   "Tank 5S Tank Vent Valve 2 Feedback - Closed" : Bool = PLC "Tank 5S Tank Vent Valve 2 Feedback - Closed" AT %I54.5, 1 s
   "RIO5_SPR_DI_54_6" : Bool = PLC RIO5_SPR_DI_54_6 AT %I54.6, 1 s
   "RIO5_SPR_DI_54_7" : Bool = PLC RIO5_SPR_DI_54_7 AT %I54.7, 1 s
   "Tank 5P BWT Level High High Switch" : Bool = PLC "Tank 5P BWT Level High High Switch" AT %I57.0, 1 s
   "RIO5 Tanks Pressure Switch Hi Hi" : Bool = PLC "RIO5 Tanks Pressure Switch Hi Hi" AT %I57.1, 1 s
   "Tank 5S BWT Level High High Switch" : Bool = PLC "Tank 5S BWT Level High High Switch" AT %I57.2, 1 s
   "RIO5_SPR_DI_57_3" : Bool = PLC RIO5_SPR_DI_57_3 AT %I57.3, 1 s
   "RIO5_SPR_DI_57_4" : Bool = PLC RIO5_SPR_DI_57_4 AT %I57.4, 1 s
   "RIO5_SPR_DI_57_5" : Bool = PLC RIO5_SPR_DI_57_5 AT %I57.5, 1 s
   "RIO5_SPR_DI_57_6" : Bool = PLC RIO5_SPR_DI_57_6 AT %I57.6, 1 s
   "RIO5_SPR_DI_57_7" : Bool = PLC RIO5_SPR_DI_57_7 AT %I57.7, 1 s
   "Tank 6P GTT Isolation Valve Feedback - Opened" : Bool = PLC "Tank 6P GTT Isolation Valve Feedback - Opened" AT %I60.0, 1 s
   "Tank 6P GTT Isolation Valve Feedback - Closed" : Bool = PLC "Tank 6P GTT Isolation Valve Feedback - Closed" AT %I60.1, 1 s
   "Tank 6P Tank Vent Valve 1 Feedback - Opened" : Bool = PLC "Tank 6P Tank Vent Valve 1 Feedback - Opened" AT %I60.2, 1 s
   "Tank 6P Tank Vent Valve 1 Feedback - Closed" : Bool = PLC "Tank 6P Tank Vent Valve 1 Feedback - Closed" AT %I60.3, 1 s
   "Tank 6P Tank Vent Valve 2 Feedback - Opened" : Bool = PLC "Tank 6P Tank Vent Valve 2 Feedback - Opened" AT %I60.4, 1 s
   "Tank 6P Tank Vent Valve 2 Feedback - Closed" : Bool = PLC "Tank 6P Tank Vent Valve 2 Feedback - Closed" AT %I60.5, 1 s
   "RIO6_SPR_DI_60_6" : Bool = PLC RIO6_SPR_DI_60_6 AT %I60.6, 1 s
   "RIO6_SPR_DI_60_7" : Bool = PLC RIO6_SPR_DI_60_7 AT %I60.7, 1 s
   "Tank 6S GTT Isolation Valve Feedback - Opened" : Bool = PLC "Tank 6S GTT Isolation Valve Feedback - Opened" AT %I63.0, 1 s
   "Tank 6S GTT Isolation Valve Feedback - Closed" : Bool = PLC "Tank 6S GTT Isolation Valve Feedback - Closed" AT %I63.1, 1 s
   "Tank 6S Tank Vent Valve 1 Feedback - Opened" : Bool = PLC "Tank 6S Tank Vent Valve 1 Feedback - Opened" AT %I63.2, 1 s
   "Tank 6S Tank Vent Valve 1 Feedback - Closed" : Bool = PLC "Tank 6S Tank Vent Valve 1 Feedback - Closed" AT %I63.3, 1 s
   "Tank 6S Tank Vent Valve 2 Feedback - Opened" : Bool = PLC "Tank 6S Tank Vent Valve 2 Feedback - Opened" AT %I63.4, 1 s
   "Tank 6S Tank Vent Valve 2 Feedback - Closed" : Bool = PLC "Tank 6S Tank Vent Valve 2 Feedback - Closed" AT %I63.5, 1 s
   "RIO6_SPR_DI_63_6" : Bool = PLC RIO6_SPR_DI_63_6 AT %I63.6, 1 s
   "RIO6_SPR_DI_63_7" : Bool = PLC RIO6_SPR_DI_63_7 AT %I63.7, 1 s
   "Tank 6P BWT Level High High Switch" : Bool = PLC "Tank 6P BWT Level High High Switch" AT %I66.0, 1 s
   "RIO6 Tanks Pressure Switch Hi Hi" : Bool = PLC "RIO6 Tanks Pressure Switch Hi Hi" AT %I66.1, 1 s
   "Tank 6S BWT Level High High Switch" : Bool = PLC "Tank 6S BWT Level High High Switch" AT %I66.2, 1 s
   "RIO6_SPR_DI_66_3" : Bool = PLC RIO6_SPR_DI_66_3 AT %I66.3, 1 s
   "RIO6_SPR_DI_66_4" : Bool = PLC RIO6_SPR_DI_66_4 AT %I66.4, 1 s
   "RIO6_SPR_DI_66_5" : Bool = PLC RIO6_SPR_DI_66_5 AT %I66.5, 1 s
   "RIO6_SPR_DI_66_7" : Bool = PLC RIO6_SPR_DI_66_7 AT %I66.7, 1 s
   "RIO6_SPR_DI_66_6" : Bool = PLC RIO6_SPR_DI_66_6 AT %I66.6, 1 s
   "APT GTT Isolation Valve Feedback - Opened" : Bool = PLC "APT GTT Isolation Valve Feedback - Opened" AT %I75.0, 1 s
   "APT GTT Isolation Valve Feedback - Closed" : Bool = PLC "APT GTT Isolation Valve Feedback - Closed" AT %I75.1, 1 s
   "APT Tank Vent Valve 1 Feedback - Opened" : Bool = PLC "APT Tank Vent Valve 1 Feedback - Opened" AT %I75.2, 1 s
   "APT Tank Vent Valve 1 Feedback - Closed" : Bool = PLC "APT Tank Vent Valve 1 Feedback - Closed" AT %I75.3, 1 s
   "APT Tank Vent Valve 2 Feedback - Opened" : Bool = PLC "APT Tank Vent Valve 2 Feedback - Opened" AT %I75.4, 1 s
   "APT Tank Vent Valve 2 Feedback - Closed" : Bool = PLC "APT Tank Vent Valve 2 Feedback - Closed" AT %I75.5, 1 s
   "RIO7_SPR_DI_175_6" : Bool = PLC RIO7_SPR_DI_175_6 AT %I75.6, 1 s
   "RIO7_SPR_DI_175_7" : Bool = PLC RIO7_SPR_DI_175_7 AT %I75.7, 1 s
   "APT BWT Level High High Switch" : Bool = PLC "APT BWT Level High High Switch" AT %I78.0, 1 s
   "RIO7 Tank Pressure Switch Hi Hi" : Bool = PLC "RIO7 Tank Pressure Switch Hi Hi" AT %I78.1, 1 s
   "RIO7_SPR_DI_178_2" : Bool = PLC RIO7_SPR_DI_178_2 AT %I78.2, 1 s
   "RIO7_SPR_DI_178_3" : Bool = PLC RIO7_SPR_DI_178_3 AT %I78.3, 1 s
   "RIO7_SPR_DI_178_4" : Bool = PLC RIO7_SPR_DI_178_4 AT %I78.4, 1 s
   "RIO7_SPR_DI_178_5" : Bool = PLC RIO7_SPR_DI_178_5 AT %I78.5, 1 s
   "RIO7_SPR_DI_178_6" : Bool = PLC RIO7_SPR_DI_178_6 AT %I78.6, 1 s
   "RIO7_SPR_DI_178_7" : Bool = PLC RIO7_SPR_DI_178_7 AT %I78.7, 1 s
   "IDB_E700 Alarms_VERY HIGH LEVEL VALUE (HH)" : Real = PLC "IDB_E700 Alarms"."VERY HIGH LEVEL VALUE (HH)" AT %DB701.DBD34, 1 s
   "IDB_E700 Alarms_HIGH LEVEL VALUE (H)" : Real = PLC "IDB_E700 Alarms"."HIGH LEVEL VALUE (H)" AT %DB701.DBD30, 1 s
   "IDB_E700 Alarms_LOW LEVEL VALUE (L)" : Real = PLC "IDB_E700 Alarms"."LOW LEVEL VALUE (L)" AT %DB701.DBD26, 1 s
   "IDB_E700 Alarms_VERY LOW LEVEL VALUE (LL)" : Real = PLC "IDB_E700 Alarms"."VERY LOW LEVEL VALUE (LL)" AT %DB701.DBD22, 1 s
   "IDB_E-600_VERY HIGH LEVEL VALUE (HH)" : Real = PLC "IDB_E-600"."VERY HIGH LEVEL VALUE (HH)" AT %DB600.DBD34, 1 s
   "IDB_E-600_HIGH LEVEL VALUE (H)" : Real = PLC "IDB_E-600"."HIGH LEVEL VALUE (H)" AT %DB600.DBD30, 1 s
   "IDB_E-600_LOW LEVEL VALUE (L)" : Real = PLC "IDB_E-600"."LOW LEVEL VALUE (L)" AT %DB600.DBD26, 1 s
   "IDB_E-600_VERY LOW LEVEL VALUE (LL)" : Real = PLC "IDB_E-600"."VERY LOW LEVEL VALUE (LL)" AT %DB600.DBD22, 1 s
   "IDB_PIT 204_VERY HIGH LEVEL VALUE (HH)" : Real = PLC "IDB_PIT 204"."VERY HIGH LEVEL VALUE (HH)" AT %DB724.DBD34, 1 s
   "IDB_PIT 204_HIGH LEVEL VALUE (H)" : Real = PLC "IDB_PIT 204"."HIGH LEVEL VALUE (H)" AT %DB724.DBD30, 1 s
   "IDB_PIT 204_LOW LEVEL VALUE (L)" : Real = PLC "IDB_PIT 204"."LOW LEVEL VALUE (L)" AT %DB724.DBD26, 1 s
   "IDB_PIT 204_VERY LOW LEVEL VALUE (LL)" : Real = PLC "IDB_PIT 204"."VERY LOW LEVEL VALUE (LL)" AT %DB724.DBD22, 1 s
   "TT426_4P_ALM_ANALOG_DB_VERY HIGH LEVEL VALUE (HH)" : Real = PLC TT426_4P_ALM_ANALOG_DB."VERY HIGH LEVEL VALUE (HH)" AT %DB2079.DBD34, 1 s
   "TT426_4P_ALM_ANALOG_DB_HIGH LEVEL VALUE (H)" : Real = PLC TT426_4P_ALM_ANALOG_DB."HIGH LEVEL VALUE (H)" AT %DB2079.DBD30, 1 s
   "TT426_4P_ALM_ANALOG_DB_LOW LEVEL VALUE (L)" : Real = PLC TT426_4P_ALM_ANALOG_DB."LOW LEVEL VALUE (L)" AT %DB2079.DBD26, 1 s
   "TT426_4P_ALM_ANALOG_DB_VERY LOW LEVEL VALUE (LL)" : Real = PLC TT426_4P_ALM_ANALOG_DB."VERY LOW LEVEL VALUE (LL)" AT %DB2079.DBD22, 1 s
   "FIT420_APT_ALM_ANALOG_DB_VERY HIGH LEVEL VALUE (HH)" : Real = PLC FIT420_APT_ALM_ANALOG_DB."VERY HIGH LEVEL VALUE (HH)" AT %DB2212.DBD34, 1 s
   "FIT420_APT_ALM_ANALOG_DB_HIGH LEVEL VALUE (H)" : Real = PLC FIT420_APT_ALM_ANALOG_DB."HIGH LEVEL VALUE (H)" AT %DB2212.DBD30, 1 s
   "FIT420_APT_ALM_ANALOG_DB_LOW LEVEL VALUE (L)" : Real = PLC FIT420_APT_ALM_ANALOG_DB."LOW LEVEL VALUE (L)" AT %DB2212.DBD26, 1 s
   "FIT420_APT_ALM_ANALOG_DB_VERY LOW LEVEL VALUE (LL)" : Real = PLC FIT420_APT_ALM_ANALOG_DB."VERY LOW LEVEL VALUE (LL)" AT %DB2212.DBD22, 1 s
   "FIT417_APT_ALM_ANALOG_DB_VERY HIGH LEVEL VALUE (HH)" : Real = PLC FIT417_APT_ALM_ANALOG_DB."VERY HIGH LEVEL VALUE (HH)" AT %DB2099.DBD34, 1 s
   "FIT417_APT_ALM_ANALOG_DB_HIGH LEVEL VALUE (H)" : Real = PLC FIT417_APT_ALM_ANALOG_DB."HIGH LEVEL VALUE (H)" AT %DB2099.DBD30, 1 s
   "FIT417_APT_ALM_ANALOG_DB_LOW LEVEL VALUE (L)" : Real = PLC FIT417_APT_ALM_ANALOG_DB."LOW LEVEL VALUE (L)" AT %DB2099.DBD26, 1 s
   "FIT417_APT_ALM_ANALOG_DB_VERY LOW LEVEL VALUE (LL)" : Real = PLC FIT417_APT_ALM_ANALOG_DB."VERY LOW LEVEL VALUE (LL)" AT %DB2099.DBD22, 1 s
   "FIT420_FPT_ALM_ANALOG_DB_VERY HIGH LEVEL VALUE (HH)" : Real = PLC FIT420_FPT_ALM_ANALOG_DB."VERY HIGH LEVEL VALUE (HH)" AT %DB2201.DBD34, 1 s
   "FIT420_FPT_ALM_ANALOG_DB_HIGH LEVEL VALUE (H)" : Real = PLC FIT420_FPT_ALM_ANALOG_DB."HIGH LEVEL VALUE (H)" AT %DB2201.DBD30, 1 s
   "FIT420_FPT_ALM_ANALOG_DB_LOW LEVEL VALUE (L)" : Real = PLC FIT420_FPT_ALM_ANALOG_DB."LOW LEVEL VALUE (L)" AT %DB2201.DBD26, 1 s
   "FIT420_FPT_ALM_ANALOG_DB_VERY LOW LEVEL VALUE (LL)" : Real = PLC FIT420_FPT_ALM_ANALOG_DB."VERY LOW LEVEL VALUE (LL)" AT %DB2201.DBD22, 1 s
   "FIT420_6S_ALM_ANALOG_DB_VERY HIGH LEVEL VALUE (HH)" : Real = PLC FIT420_6S_ALM_ANALOG_DB."VERY HIGH LEVEL VALUE (HH)" AT %DB2211.DBD34, 1 s
   "FIT420_6S_ALM_ANALOG_DB_HIGH LEVEL VALUE (H)" : Real = PLC FIT420_6S_ALM_ANALOG_DB."HIGH LEVEL VALUE (H)" AT %DB2211.DBD30, 1 s
   "FIT420_6S_ALM_ANALOG_DB_LOW LEVEL VALUE (L)" : Real = PLC FIT420_6S_ALM_ANALOG_DB."LOW LEVEL VALUE (L)" AT %DB2211.DBD26, 1 s
   "FIT420_6S_ALM_ANALOG_DB_VERY LOW LEVEL VALUE (LL)" : Real = PLC FIT420_6S_ALM_ANALOG_DB."VERY LOW LEVEL VALUE (LL)" AT %DB2211.DBD22, 1 s
   "FIT417_6S_ALM_ANALOG_DB_VERY HIGH LEVEL VALUE (HH)" : Real = PLC FIT417_6S_ALM_ANALOG_DB."VERY HIGH LEVEL VALUE (HH)" AT %DB2098.DBD34, 1 s
   "FIT417_6S_ALM_ANALOG_DB_HIGH LEVEL VALUE (H)" : Real = PLC FIT417_6S_ALM_ANALOG_DB."HIGH LEVEL VALUE (H)" AT %DB2098.DBD30, 1 s
   "FIT417_6S_ALM_ANALOG_DB_LOW LEVEL VALUE (L)" : Real = PLC FIT417_6S_ALM_ANALOG_DB."LOW LEVEL VALUE (L)" AT %DB2098.DBD26, 1 s
   "FIT417_6S_ALM_ANALOG_DB_VERY LOW LEVEL VALUE (LL)" : Real = PLC FIT417_6S_ALM_ANALOG_DB."VERY LOW LEVEL VALUE (LL)" AT %DB2098.DBD22, 1 s
   "FIT420_6P_ALM_ANALOG_DB_VERY HIGH LEVEL VALUE (HH)" : Real = PLC FIT420_6P_ALM_ANALOG_DB."VERY HIGH LEVEL VALUE (HH)" AT %DB2210.DBD34, 1 s
   "FIT420_6P_ALM_ANALOG_DB_HIGH LEVEL VALUE (H)" : Real = PLC FIT420_6P_ALM_ANALOG_DB."HIGH LEVEL VALUE (H)" AT %DB2210.DBD30, 1 s
   "FIT420_6P_ALM_ANALOG_DB_LOW LEVEL VALUE (L)" : Real = PLC FIT420_6P_ALM_ANALOG_DB."LOW LEVEL VALUE (L)" AT %DB2210.DBD26, 1 s
   "FIT420_6P_ALM_ANALOG_DB_VERY LOW LEVEL VALUE (LL)" : Real = PLC FIT420_6P_ALM_ANALOG_DB."VERY LOW LEVEL VALUE (LL)" AT %DB2210.DBD22, 1 s
   "FIT418_6P__ALM_ANALOG_DB_VERY HIGH LEVEL VALUE (HH)" : Real = PLC "FIT418_6P__ALM_ANALOG_DB"."VERY HIGH LEVEL VALUE (HH)" AT %DB2097.DBD34, 1 s
   "FIT418_6P__ALM_ANALOG_DB_HIGH LEVEL VALUE (H)" : Real = PLC "FIT418_6P__ALM_ANALOG_DB"."HIGH LEVEL VALUE (H)" AT %DB2097.DBD30, 1 s
   "FIT418_6P__ALM_ANALOG_DB_LOW LEVEL VALUE (L)" : Real = PLC "FIT418_6P__ALM_ANALOG_DB"."LOW LEVEL VALUE (L)" AT %DB2097.DBD26, 1 s
   "FIT418_6P__ALM_ANALOG_DB_VERY LOW LEVEL VALUE (LL)" : Real = PLC "FIT418_6P__ALM_ANALOG_DB"."VERY LOW LEVEL VALUE (LL)" AT %DB2097.DBD22, 1 s
   "FIT420_5S_ALM_ANALOG_DB_VERY HIGH LEVEL VALUE (HH)" : Real = PLC FIT420_5S_ALM_ANALOG_DB."VERY HIGH LEVEL VALUE (HH)" AT %DB2209.DBD34, 1 s
   "FIT420_5S_ALM_ANALOG_DB_HIGH LEVEL VALUE (H)" : Real = PLC FIT420_5S_ALM_ANALOG_DB."HIGH LEVEL VALUE (H)" AT %DB2209.DBD30, 1 s
   "FIT420_5S_ALM_ANALOG_DB_LOW LEVEL VALUE (L)" : Real = PLC FIT420_5S_ALM_ANALOG_DB."LOW LEVEL VALUE (L)" AT %DB2209.DBD26, 1 s
   "FIT420_5S_ALM_ANALOG_DB_VERY LOW LEVEL VALUE (LL)" : Real = PLC FIT420_5S_ALM_ANALOG_DB."VERY LOW LEVEL VALUE (LL)" AT %DB2209.DBD22, 1 s
   "FIT417_5S_ALM_ANALOG_DB_VERY HIGH LEVEL VALUE (HH)" : Real = PLC FIT417_5S_ALM_ANALOG_DB."VERY HIGH LEVEL VALUE (HH)" AT %DB2096.DBD34, 1 s
   "FIT417_5S_ALM_ANALOG_DB_HIGH LEVEL VALUE (H)" : Real = PLC FIT417_5S_ALM_ANALOG_DB."HIGH LEVEL VALUE (H)" AT %DB2096.DBD30, 1 s
   "FIT417_5S_ALM_ANALOG_DB_LOW LEVEL VALUE (L)" : Real = PLC FIT417_5S_ALM_ANALOG_DB."LOW LEVEL VALUE (L)" AT %DB2096.DBD26, 1 s
   "FIT417_5S_ALM_ANALOG_DB_VERY LOW LEVEL VALUE (LL)" : Real = PLC FIT417_5S_ALM_ANALOG_DB."VERY LOW LEVEL VALUE (LL)" AT %DB2096.DBD22, 1 s
   "FIT418_5P__ALM_ANALOG_DB_VERY HIGH LEVEL VALUE (HH)" : Real = PLC "FIT418_5P__ALM_ANALOG_DB"."VERY HIGH LEVEL VALUE (HH)" AT %DB2095.DBD34, 1 s
   "FIT418_5P__ALM_ANALOG_DB_HIGH LEVEL VALUE (H)" : Real = PLC "FIT418_5P__ALM_ANALOG_DB"."HIGH LEVEL VALUE (H)" AT %DB2095.DBD30, 1 s
   "FIT418_5P__ALM_ANALOG_DB_LOW LEVEL VALUE (L)" : Real = PLC "FIT418_5P__ALM_ANALOG_DB"."LOW LEVEL VALUE (L)" AT %DB2095.DBD26, 1 s
   "FIT418_5P__ALM_ANALOG_DB_VERY LOW LEVEL VALUE (LL)" : Real = PLC "FIT418_5P__ALM_ANALOG_DB"."VERY LOW LEVEL VALUE (LL)" AT %DB2095.DBD22, 1 s
   "FIT420_5P_ALM_ANALOG_DB_VERY HIGH LEVEL VALUE (HH)" : Real = PLC FIT420_5P_ALM_ANALOG_DB."VERY HIGH LEVEL VALUE (HH)" AT %DB2208.DBD34, 1 s
   "FIT420_5P_ALM_ANALOG_DB_HIGH LEVEL VALUE (H)" : Real = PLC FIT420_5P_ALM_ANALOG_DB."HIGH LEVEL VALUE (H)" AT %DB2208.DBD30, 1 s
   "FIT420_5P_ALM_ANALOG_DB_LOW LEVEL VALUE (L)" : Real = PLC FIT420_5P_ALM_ANALOG_DB."LOW LEVEL VALUE (L)" AT %DB2208.DBD26, 1 s
   "FIT420_5P_ALM_ANALOG_DB_VERY LOW LEVEL VALUE (LL)" : Real = PLC FIT420_5P_ALM_ANALOG_DB."VERY LOW LEVEL VALUE (LL)" AT %DB2208.DBD22, 1 s
   "FIT420_4S_ALM_ANALOG_DB_VERY HIGH LEVEL VALUE (HH)" : Real = PLC FIT420_4S_ALM_ANALOG_DB."VERY HIGH LEVEL VALUE (HH)" AT %DB2207.DBD34, 1 s
   "FIT420_4S_ALM_ANALOG_DB_HIGH LEVEL VALUE (H)" : Real = PLC FIT420_4S_ALM_ANALOG_DB."HIGH LEVEL VALUE (H)" AT %DB2207.DBD30, 1 s
   "FIT420_4S_ALM_ANALOG_DB_LOW LEVEL VALUE (L)" : Real = PLC FIT420_4S_ALM_ANALOG_DB."LOW LEVEL VALUE (L)" AT %DB2207.DBD26, 1 s
   "FIT420_4S_ALM_ANALOG_DB_VERY LOW LEVEL VALUE (LL)" : Real = PLC FIT420_4S_ALM_ANALOG_DB."VERY LOW LEVEL VALUE (LL)" AT %DB2207.DBD22, 1 s
   "FIT417_4S_ALM_ANALOG_DB_VERY HIGH LEVEL VALUE (HH)" : Real = PLC FIT417_4S_ALM_ANALOG_DB."VERY HIGH LEVEL VALUE (HH)" AT %DB2094.DBD34, 1 s
   "FIT417_4S_ALM_ANALOG_DB_HIGH LEVEL VALUE (H)" : Real = PLC FIT417_4S_ALM_ANALOG_DB."HIGH LEVEL VALUE (H)" AT %DB2094.DBD30, 1 s
   "FIT417_4S_ALM_ANALOG_DB_LOW LEVEL VALUE (L)" : Real = PLC FIT417_4S_ALM_ANALOG_DB."LOW LEVEL VALUE (L)" AT %DB2094.DBD26, 1 s
   "FIT417_4S_ALM_ANALOG_DB_VERY LOW LEVEL VALUE (LL)" : Real = PLC FIT417_4S_ALM_ANALOG_DB."VERY LOW LEVEL VALUE (LL)" AT %DB2094.DBD22, 1 s
   "LT422 4P  TANK LEVEL ALARM_VERY HIGH LEVEL VALUE (HH)" : Real = PLC "LT422 4P  TANK LEVEL ALARM"."VERY HIGH LEVEL VALUE (HH)" AT %DB2233.DBD34, 1 s
   "LT422 4P  TANK LEVEL ALARM_HIGH LEVEL VALUE (H)" : Real = PLC "LT422 4P  TANK LEVEL ALARM"."HIGH LEVEL VALUE (H)" AT %DB2233.DBD30, 1 s
   "LT422 4P  TANK LEVEL ALARM_LOW LEVEL VALUE (L)" : Real = PLC "LT422 4P  TANK LEVEL ALARM"."LOW LEVEL VALUE (L)" AT %DB2233.DBD26, 1 s
   "LT422 4P  TANK LEVEL ALARM_VERY LOW LEVEL VALUE (LL)" : Real = PLC "LT422 4P  TANK LEVEL ALARM"."VERY LOW LEVEL VALUE (LL)" AT %DB2233.DBD22, 1 s
   "FIT420_4P_ALM_ANALOG_DB_VERY HIGH LEVEL VALUE (HH)" : Real = PLC FIT420_4P_ALM_ANALOG_DB."VERY HIGH LEVEL VALUE (HH)" AT %DB2206.DBD34, 1 s
   "FIT420_4P_ALM_ANALOG_DB_HIGH LEVEL VALUE (H)" : Real = PLC FIT420_4P_ALM_ANALOG_DB."HIGH LEVEL VALUE (H)" AT %DB2206.DBD30, 1 s
   "FIT420_4P_ALM_ANALOG_DB_LOW LEVEL VALUE (L)" : Real = PLC FIT420_4P_ALM_ANALOG_DB."LOW LEVEL VALUE (L)" AT %DB2206.DBD26, 1 s
   "FIT420_4P_ALM_ANALOG_DB_VERY LOW LEVEL VALUE (LL)" : Real = PLC FIT420_4P_ALM_ANALOG_DB."VERY LOW LEVEL VALUE (LL)" AT %DB2206.DBD22, 1 s
   "FIT418_4P__ALM_ANALOG_DB_VERY HIGH LEVEL VALUE (HH)" : Real = PLC "FIT418_4P__ALM_ANALOG_DB"."VERY HIGH LEVEL VALUE (HH)" AT %DB2093.DBD34, 1 s
   "FIT418_4P__ALM_ANALOG_DB_HIGH LEVEL VALUE (H)" : Real = PLC "FIT418_4P__ALM_ANALOG_DB"."HIGH LEVEL VALUE (H)" AT %DB2093.DBD30, 1 s
   "FIT418_4P__ALM_ANALOG_DB_LOW LEVEL VALUE (L)" : Real = PLC "FIT418_4P__ALM_ANALOG_DB"."LOW LEVEL VALUE (L)" AT %DB2093.DBD26, 1 s
   "FIT418_4P__ALM_ANALOG_DB_VERY LOW LEVEL VALUE (LL)" : Real = PLC "FIT418_4P__ALM_ANALOG_DB"."VERY LOW LEVEL VALUE (LL)" AT %DB2093.DBD22, 1 s
   "FIT420_3S_ALM_ANALOG_DB_VERY HIGH LEVEL VALUE (HH)" : Real = PLC FIT420_3S_ALM_ANALOG_DB."VERY HIGH LEVEL VALUE (HH)" AT %DB2205.DBD34, 1 s
   "FIT420_3S_ALM_ANALOG_DB_HIGH LEVEL VALUE (H)" : Real = PLC FIT420_3S_ALM_ANALOG_DB."HIGH LEVEL VALUE (H)" AT %DB2205.DBD30, 1 s
   "FIT420_3S_ALM_ANALOG_DB_LOW LEVEL VALUE (L)" : Real = PLC FIT420_3S_ALM_ANALOG_DB."LOW LEVEL VALUE (L)" AT %DB2205.DBD26, 1 s
   "FIT420_3S_ALM_ANALOG_DB_VERY LOW LEVEL VALUE (LL)" : Real = PLC FIT420_3S_ALM_ANALOG_DB."VERY LOW LEVEL VALUE (LL)" AT %DB2205.DBD22, 1 s
   "FIT417_3S_ALM_ANALOG_DB_VERY HIGH LEVEL VALUE (HH)" : Real = PLC FIT417_3S_ALM_ANALOG_DB."VERY HIGH LEVEL VALUE (HH)" AT %DB2092.DBD34, 1 s
   "FIT417_3S_ALM_ANALOG_DB_HIGH LEVEL VALUE (H)" : Real = PLC FIT417_3S_ALM_ANALOG_DB."HIGH LEVEL VALUE (H)" AT %DB2092.DBD30, 1 s
   "FIT417_3S_ALM_ANALOG_DB_LOW LEVEL VALUE (L)" : Real = PLC FIT417_3S_ALM_ANALOG_DB."LOW LEVEL VALUE (L)" AT %DB2092.DBD26, 1 s
   "FIT417_3S_ALM_ANALOG_DB_VERY LOW LEVEL VALUE (LL)" : Real = PLC FIT417_3S_ALM_ANALOG_DB."VERY LOW LEVEL VALUE (LL)" AT %DB2092.DBD22, 1 s
   "FIT418_3P__ALM_ANALOG_DB_VERY HIGH LEVEL VALUE (HH)" : Real = PLC "FIT418_3P__ALM_ANALOG_DB"."VERY HIGH LEVEL VALUE (HH)" AT %DB2091.DBD34, 1 s
   "FIT418_3P__ALM_ANALOG_DB_HIGH LEVEL VALUE (H)" : Real = PLC "FIT418_3P__ALM_ANALOG_DB"."HIGH LEVEL VALUE (H)" AT %DB2091.DBD30, 1 s
   "FIT418_3P__ALM_ANALOG_DB_LOW LEVEL VALUE (L)" : Real = PLC "FIT418_3P__ALM_ANALOG_DB"."LOW LEVEL VALUE (L)" AT %DB2091.DBD26, 1 s
   "FIT418_3P__ALM_ANALOG_DB_VERY LOW LEVEL VALUE (LL)" : Real = PLC "FIT418_3P__ALM_ANALOG_DB"."VERY LOW LEVEL VALUE (LL)" AT %DB2091.DBD22, 1 s
   "FIT420_3P_ALM_ANALOG_DB_VERY HIGH LEVEL VALUE (HH)" : Real = PLC FIT420_3P_ALM_ANALOG_DB."VERY HIGH LEVEL VALUE (HH)" AT %DB2204.DBD34, 1 s
   "FIT420_3P_ALM_ANALOG_DB_HIGH LEVEL VALUE (H)" : Real = PLC FIT420_3P_ALM_ANALOG_DB."HIGH LEVEL VALUE (H)" AT %DB2204.DBD30, 1 s
   "FIT420_3P_ALM_ANALOG_DB_LOW LEVEL VALUE (L)" : Real = PLC FIT420_3P_ALM_ANALOG_DB."LOW LEVEL VALUE (L)" AT %DB2204.DBD26, 1 s
   "FIT420_3P_ALM_ANALOG_DB_VERY LOW LEVEL VALUE (LL)" : Real = PLC FIT420_3P_ALM_ANALOG_DB."VERY LOW LEVEL VALUE (LL)" AT %DB2204.DBD22, 1 s
   "FIT420_1S_ALM_ANALOG_DB_VERY HIGH LEVEL VALUE (HH)" : Real = PLC FIT420_1S_ALM_ANALOG_DB."VERY HIGH LEVEL VALUE (HH)" AT %DB2203.DBD34, 1 s
   "FIT420_1S_ALM_ANALOG_DB_HIGH LEVEL VALUE (H)" : Real = PLC FIT420_1S_ALM_ANALOG_DB."HIGH LEVEL VALUE (H)" AT %DB2203.DBD30, 1 s
   "FIT420_1S_ALM_ANALOG_DB_LOW LEVEL VALUE (L)" : Real = PLC FIT420_1S_ALM_ANALOG_DB."LOW LEVEL VALUE (L)" AT %DB2203.DBD26, 1 s
   "FIT420_1S_ALM_ANALOG_DB_VERY LOW LEVEL VALUE (LL)" : Real = PLC FIT420_1S_ALM_ANALOG_DB."VERY LOW LEVEL VALUE (LL)" AT %DB2203.DBD22, 1 s
   "FIT417_1S__ALM_ANALOG_DB_VERY HIGH LEVEL VALUE (HH)" : Real = PLC "FIT417_1S__ALM_ANALOG_DB"."VERY HIGH LEVEL VALUE (HH)" AT %DB2090.DBD34, 1 s
   "FIT417_1S__ALM_ANALOG_DB_HIGH LEVEL VALUE (H)" : Real = PLC "FIT417_1S__ALM_ANALOG_DB"."HIGH LEVEL VALUE (H)" AT %DB2090.DBD30, 1 s
   "FIT417_1S__ALM_ANALOG_DB_LOW LEVEL VALUE (L)" : Real = PLC "FIT417_1S__ALM_ANALOG_DB"."LOW LEVEL VALUE (L)" AT %DB2090.DBD26, 1 s
   "FIT417_1S__ALM_ANALOG_DB_VERY LOW LEVEL VALUE (LL)" : Real = PLC "FIT417_1S__ALM_ANALOG_DB"."VERY LOW LEVEL VALUE (LL)" AT %DB2090.DBD22, 1 s
   "FIT420_1P_ALM_ANALOG_DB_VERY HIGH LEVEL VALUE (HH)" : Real = PLC FIT420_1P_ALM_ANALOG_DB."VERY HIGH LEVEL VALUE (HH)" AT %DB2202.DBD34, 1 s
   "FIT420_1P_ALM_ANALOG_DB_HIGH LEVEL VALUE (H)" : Real = PLC FIT420_1P_ALM_ANALOG_DB."HIGH LEVEL VALUE (H)" AT %DB2202.DBD30, 1 s
   "FIT420_1P_ALM_ANALOG_DB_LOW LEVEL VALUE (L)" : Real = PLC FIT420_1P_ALM_ANALOG_DB."LOW LEVEL VALUE (L)" AT %DB2202.DBD26, 1 s
   "FIT420_1P_ALM_ANALOG_DB_VERY LOW LEVEL VALUE (LL)" : Real = PLC FIT420_1P_ALM_ANALOG_DB."VERY LOW LEVEL VALUE (LL)" AT %DB2202.DBD22, 1 s
   "FIT418_1P__ALM_ANALOG_DB_VERY HIGH LEVEL VALUE (HH)" : Real = PLC "FIT418_1P__ALM_ANALOG_DB"."VERY HIGH LEVEL VALUE (HH)" AT %DB2089.DBD34, 1 s
   "FIT418_1P__ALM_ANALOG_DB_HIGH LEVEL VALUE (H)" : Real = PLC "FIT418_1P__ALM_ANALOG_DB"."HIGH LEVEL VALUE (H)" AT %DB2089.DBD30, 1 s
   "FIT418_1P__ALM_ANALOG_DB_LOW LEVEL VALUE (L)" : Real = PLC "FIT418_1P__ALM_ANALOG_DB"."LOW LEVEL VALUE (L)" AT %DB2089.DBD26, 1 s
   "FIT418_1P__ALM_ANALOG_DB_VERY LOW LEVEL VALUE (LL)" : Real = PLC "FIT418_1P__ALM_ANALOG_DB"."VERY LOW LEVEL VALUE (LL)" AT %DB2089.DBD22, 1 s
   "FIT418_FPT__ALM_ANALOG_DB_VERY HIGH LEVEL VALUE (HH)" : Real = PLC "FIT418_FPT__ALM_ANALOG_DB"."VERY HIGH LEVEL VALUE (HH)" AT %DB2088.DBD34, 1 s
   "FIT418_FPT__ALM_ANALOG_DB_HIGH LEVEL VALUE (H)" : Real = PLC "FIT418_FPT__ALM_ANALOG_DB"."HIGH LEVEL VALUE (H)" AT %DB2088.DBD30, 1 s
   "FIT418_FPT__ALM_ANALOG_DB_LOW LEVEL VALUE (L)" : Real = PLC "FIT418_FPT__ALM_ANALOG_DB"."LOW LEVEL VALUE (L)" AT %DB2088.DBD26, 1 s
   "FIT418_FPT__ALM_ANALOG_DB_VERY LOW LEVEL VALUE (LL)" : Real = PLC "FIT418_FPT__ALM_ANALOG_DB"."VERY LOW LEVEL VALUE (LL)" AT %DB2088.DBD22, 1 s
   "TT426_1P_ALM_ANALOG_DB_VERY HIGH LEVEL VALUE (HH)" : Real = PLC TT426_1P_ALM_ANALOG_DB."VERY HIGH LEVEL VALUE (HH)" AT %DB2075.DBD34, 1 s
   "TT426_1P_ALM_ANALOG_DB_HIGH LEVEL VALUE (H)" : Real = PLC TT426_1P_ALM_ANALOG_DB."HIGH LEVEL VALUE (H)" AT %DB2075.DBD30, 1 s
   "TT426_1P_ALM_ANALOG_DB_LOW LEVEL VALUE (L)" : Real = PLC TT426_1P_ALM_ANALOG_DB."LOW LEVEL VALUE (L)" AT %DB2075.DBD26, 1 s
   "TT426_1P_ALM_ANALOG_DB_VERY LOW LEVEL VALUE (LL)" : Real = PLC TT426_1P_ALM_ANALOG_DB."VERY LOW LEVEL VALUE (LL)" AT %DB2075.DBD22, 1 s
   "PIT424_RIO1_ALM_ANALOG_DB_VERY HIGH LEVEL VALUE (HH)" : Real = PLC PIT424_RIO1_ALM_ANALOG_DB."VERY HIGH LEVEL VALUE (HH)" AT %DB2219.DBD34, 1 s
   "PIT424_RIO1_ALM_ANALOG_DB_HIGH LEVEL VALUE (H)" : Real = PLC PIT424_RIO1_ALM_ANALOG_DB."HIGH LEVEL VALUE (H)" AT %DB2219.DBD30, 1 s
   "PIT424_RIO1_ALM_ANALOG_DB_LOW LEVEL VALUE (L)" : Real = PLC PIT424_RIO1_ALM_ANALOG_DB."LOW LEVEL VALUE (L)" AT %DB2219.DBD26, 1 s
   "PIT424_RIO1_ALM_ANALOG_DB_VERY LOW LEVEL VALUE (LL)" : Real = PLC PIT424_RIO1_ALM_ANALOG_DB."VERY LOW LEVEL VALUE (LL)" AT %DB2219.DBD22, 1 s
   "TT426_1S_ALM_ANALOG_DB_VERY HIGH LEVEL VALUE (HH)" : Real = PLC TT426_1S_ALM_ANALOG_DB."VERY HIGH LEVEL VALUE (HH)" AT %DB2076.DBD34, 1 s
   "TT426_1S_ALM_ANALOG_DB_HIGH LEVEL VALUE (H)" : Real = PLC TT426_1S_ALM_ANALOG_DB."HIGH LEVEL VALUE (H)" AT %DB2076.DBD30, 1 s
   "TT426_1S_ALM_ANALOG_DB_LOW LEVEL VALUE (L)" : Real = PLC TT426_1S_ALM_ANALOG_DB."LOW LEVEL VALUE (L)" AT %DB2076.DBD26, 1 s
   "TT426_1S_ALM_ANALOG_DB_VERY LOW LEVEL VALUE (LL)" : Real = PLC TT426_1S_ALM_ANALOG_DB."VERY LOW LEVEL VALUE (LL)" AT %DB2076.DBD22, 1 s
   "TT426_3P_ALM_ANALOG_DB_VERY HIGH LEVEL VALUE (HH)" : Real = PLC TT426_3P_ALM_ANALOG_DB."VERY HIGH LEVEL VALUE (HH)" AT %DB2077.DBD34, 1 s
   "TT426_3P_ALM_ANALOG_DB_HIGH LEVEL VALUE (H)" : Real = PLC TT426_3P_ALM_ANALOG_DB."HIGH LEVEL VALUE (H)" AT %DB2077.DBD30, 1 s
   "TT426_3P_ALM_ANALOG_DB_LOW LEVEL VALUE (L)" : Real = PLC TT426_3P_ALM_ANALOG_DB."LOW LEVEL VALUE (L)" AT %DB2077.DBD26, 1 s
   "TT426_3P_ALM_ANALOG_DB_VERY LOW LEVEL VALUE (LL)" : Real = PLC TT426_3P_ALM_ANALOG_DB."VERY LOW LEVEL VALUE (LL)" AT %DB2077.DBD22, 1 s
   "PIT424_RIO3_ALM_ANALOG_DB_VERY HIGH LEVEL VALUE (HH)" : Real = PLC PIT424_RIO3_ALM_ANALOG_DB."VERY HIGH LEVEL VALUE (HH)" AT %DB2220.DBD34, 1 s
   "PIT424_RIO3_ALM_ANALOG_DB_HIGH LEVEL VALUE (H)" : Real = PLC PIT424_RIO3_ALM_ANALOG_DB."HIGH LEVEL VALUE (H)" AT %DB2220.DBD30, 1 s
   "PIT424_RIO3_ALM_ANALOG_DB_LOW LEVEL VALUE (L)" : Real = PLC "2102_TIME_CALCS_DB"."PRE-DWEL_Warning 1" AT %DB2220.DBD26, 1 s
   "PIT424_RIO3_ALM_ANALOG_DB_VERY LOW LEVEL VALUE (LL)" : Real = PLC PIT424_RIO3_ALM_ANALOG_DB."VERY LOW LEVEL VALUE (LL)" AT %DB2220.DBD22, 1 s
   "TT426_3S_ALM_ANALOG_DB_VERY HIGH LEVEL VALUE (HH)" : Real = PLC TT426_3S_ALM_ANALOG_DB."VERY HIGH LEVEL VALUE (HH)" AT %DB2078.DBD34, 1 s
   "TT426_3S_ALM_ANALOG_DB_HIGH LEVEL VALUE (H)" : Real = PLC TT426_3S_ALM_ANALOG_DB."HIGH LEVEL VALUE (H)" AT %DB2078.DBD30, 1 s
   "TT426_3S_ALM_ANALOG_DB_LOW LEVEL VALUE (L)" : Real = PLC TT426_3S_ALM_ANALOG_DB."LOW LEVEL VALUE (L)" AT %DB2078.DBD26, 1 s
   "TT426_3S_ALM_ANALOG_DB_VERY LOW LEVEL VALUE (LL)" : Real = PLC TT426_3S_ALM_ANALOG_DB."VERY LOW LEVEL VALUE (LL)" AT %DB2078.DBD22, 1 s
   "PIT424_RIO4_ALM_ANALOG_DB_VERY HIGH LEVEL VALUE (HH)" : Real = PLC PIT424_RIO4_ALM_ANALOG_DB."VERY HIGH LEVEL VALUE (HH)" AT %DB2221.DBD34, 1 s
   "PIT424_RIO4_ALM_ANALOG_DB_HIGH LEVEL VALUE (H)" : Real = PLC PIT424_RIO4_ALM_ANALOG_DB."HIGH LEVEL VALUE (H)" AT %DB2221.DBD30, 1 s
   "PIT424_RIO4_ALM_ANALOG_DB_LOW LEVEL VALUE (L)" : Real = PLC PIT424_RIO4_ALM_ANALOG_DB."LOW LEVEL VALUE (L)" AT %DB2221.DBD26, 1 s
   "PIT424_RIO4_ALM_ANALOG_DB_VERY LOW LEVEL VALUE (LL)" : Real = PLC PIT424_RIO4_ALM_ANALOG_DB."VERY LOW LEVEL VALUE (LL)" AT %DB2221.DBD22, 1 s
   "TT426_FPT_ALM_ANALOG_DB_VERY HIGH LEVEL VALUE (HH)" : Real = PLC TT426_FPT_ALM_ANALOG_DB."VERY HIGH LEVEL VALUE (HH)" AT %DB2074.DBD34, 1 s
   "TT426_FPT_ALM_ANALOG_DB_HIGH LEVEL VALUE (H)" : Real = PLC TT426_FPT_ALM_ANALOG_DB."HIGH LEVEL VALUE (H)" AT %DB2074.DBD30, 1 s
   "TT426_FPT_ALM_ANALOG_DB_LOW LEVEL VALUE (L)" : Real = PLC TT426_FPT_ALM_ANALOG_DB."LOW LEVEL VALUE (L)" AT %DB2074.DBD26, 1 s
   "TT426_FPT_ALM_ANALOG_DB_VERY LOW LEVEL VALUE (LL)" : Real = PLC TT426_FPT_ALM_ANALOG_DB."VERY LOW LEVEL VALUE (LL)" AT %DB2074.DBD22, 1 s
   "PT415_RIO4_ALM_ANALOG_DB_VERY HIGH LEVEL VALUE (HH)" : Real = PLC PT415_RIO4_ALM_ANALOG_DB."VERY HIGH LEVEL VALUE (HH)" AT %DB2216.DBD34, 1 s
   "PT415_RIO4_ALM_ANALOG_DB_HIGH LEVEL VALUE (H)" : Real = PLC "2086_Times".DEOX_PRE_GTT_CLS_DLY AT %DB2216.DBD30, 1 s
   "PT415_RIO4_ALM_ANALOG_DB_LOW LEVEL VALUE (L)" : Real = PLC PT415_RIO4_ALM_ANALOG_DB."LOW LEVEL VALUE (L)" AT %DB2216.DBD26, 1 s
   "PT415_RIO4_ALM_ANALOG_DB_VERY LOW LEVEL VALUE (LL)" : Real = PLC PT415_RIO4_ALM_ANALOG_DB."VERY LOW LEVEL VALUE (LL)" AT %DB2216.DBD22, 1 s
   "PIT353_ALM_ANALOG_DB72_VERY HIGH LEVEL VALUE (HH)" : Real = PLC PIT353_ALM_ANALOG_DB72."VERY HIGH LEVEL VALUE (HH)" AT %DB72.DBD34, 1 s
   "PIT353_ALM_ANALOG_DB72_HIGH LEVEL VALUE (H)" : Real = PLC PIT353_ALM_ANALOG_DB72."HIGH LEVEL VALUE (H)" AT %DB72.DBD30, 1 s
   "PIT353_ALM_ANALOG_DB72_LOW LEVEL VALUE (L)" : Real = PLC PIT353_ALM_ANALOG_DB72."LOW LEVEL VALUE (L)" AT %DB72.DBD26, 1 s
   "PIT353_ALM_ANALOG_DB72_VERY LOW LEVEL VALUE (LL)" : Real = PLC PIT353_ALM_ANALOG_DB72."VERY LOW LEVEL VALUE (LL)" AT %DB72.DBD22, 1 s
   "TIT408_ALM_ANALOG_DB75_VERY HIGH LEVEL VALUE (HH)" : Real = PLC TIT408_ALM_ANALOG_DB75."VERY HIGH LEVEL VALUE (HH)" AT %DB75.DBD34, 1 s
   "TIT408_ALM_ANALOG_DB75_HIGH LEVEL VALUE (H)" : Real = PLC TIT408_ALM_ANALOG_DB75."HIGH LEVEL VALUE (H)" AT %DB75.DBD30, 1 s
   "TIT408_ALM_ANALOG_DB75_LOW LEVEL VALUE (L)" : Real = PLC TIT408_ALM_ANALOG_DB75."LOW LEVEL VALUE (L)" AT %DB75.DBD26, 1 s
   "TIT408_ALM_ANALOG_DB75_VERY LOW LEVEL VALUE (LL)" : Real = PLC TIT408_ALM_ANALOG_DB75."VERY LOW LEVEL VALUE (LL)" AT %DB75.DBD22, 1 s
   "PIT348_ALM_ANALOG_DB73_VERY HIGH LEVEL VALUE (HH)" : Real = PLC PIT348_ALM_ANALOG_DB73."VERY HIGH LEVEL VALUE (HH)" AT %DB73.DBD34, 1 s
   "PIT348_ALM_ANALOG_DB73_HIGH LEVEL VALUE (H)" : Real = PLC PIT348_ALM_ANALOG_DB73."HIGH LEVEL VALUE (H)" AT %DB73.DBD30, 1 s
   "PIT348_ALM_ANALOG_DB73_LOW LEVEL VALUE (L)" : Real = PLC PIT348_ALM_ANALOG_DB73."LOW LEVEL VALUE (L)" AT %DB73.DBD26, 1 s
   "PIT348_ALM_ANALOG_DB73_VERY LOW LEVEL VALUE (LL)" : Real = PLC PIT348_ALM_ANALOG_DB73."VERY LOW LEVEL VALUE (LL)" AT %DB73.DBD22, 1 s
   "PIT358_ALM_ANALOG_DB78_VERY HIGH LEVEL VALUE (HH)" : Real = PLC PIT358_ALM_ANALOG_DB78."VERY HIGH LEVEL VALUE (HH)" AT %DB78.DBD34, 1 s
   "PIT358_ALM_ANALOG_DB78_HIGH LEVEL VALUE (H)" : Real = PLC PIT358_ALM_ANALOG_DB78."HIGH LEVEL VALUE (H)" AT %DB78.DBD30, 1 s
   "PIT358_ALM_ANALOG_DB78_LOW LEVEL VALUE (L)" : Real = PLC PIT358_ALM_ANALOG_DB78."LOW LEVEL VALUE (L)" AT %DB78.DBD26, 1 s
   "PIT358_ALM_ANALOG_DB78_VERY LOW LEVEL VALUE (LL)" : Real = PLC PIT358_ALM_ANALOG_DB78."VERY LOW LEVEL VALUE (LL)" AT %DB78.DBD22, 1 s
   "TT002_ALM_ANALOG_DB76_VERY HIGH LEVEL VALUE (HH)" : Real = PLC TT002_ALM_ANALOG_DB76."VERY HIGH LEVEL VALUE (HH)" AT %DB76.DBD34, 1 s
   "TT002_ALM_ANALOG_DB76_HIGH LEVEL VALUE (H)" : Real = PLC TT002_ALM_ANALOG_DB76."HIGH LEVEL VALUE (H)" AT %DB76.DBD30, 1 s
   "TT002_ALM_ANALOG_DB76_LOW LEVEL VALUE (L)" : Real = PLC TT002_ALM_ANALOG_DB76."LOW LEVEL VALUE (L)" AT %DB76.DBD26, 1 s
   "TT002_ALM_ANALOG_DB76_VERY LOW LEVEL VALUE (LL)" : Real = PLC TT002_ALM_ANALOG_DB76."VERY LOW LEVEL VALUE (LL)" AT %DB76.DBD22, 1 s
   "PT415PORT_ALM_ANALOG_DB_VERY HIGH LEVEL VALUE (HH)" : Real = PLC PT415PORT_ALM_ANALOG_DB."VERY HIGH LEVEL VALUE (HH)" AT %DB2069.DBD34, 1 s
   "PT415PORT_ALM_ANALOG_DB_HIGH LEVEL VALUE (H)" : Real = PLC PT415PORT_ALM_ANALOG_DB."HIGH LEVEL VALUE (H)" AT %DB2069.DBD30, 1 s
   "PT415PORT_ALM_ANALOG_DB_LOW LEVEL VALUE (L)" : Real = PLC PT415PORT_ALM_ANALOG_DB."LOW LEVEL VALUE (L)" AT %DB2069.DBD26, 1 s
   "PT415PORT_ALM_ANALOG_DB_VERY LOW LEVEL VALUE (LL)" : Real = PLC PT415PORT_ALM_ANALOG_DB."VERY LOW LEVEL VALUE (LL)" AT %DB2069.DBD22, 1 s
   "502_ALM_ANALOG_IDB PIT 416_VERY HIGH LEVEL VALUE (HH)" : Real = PLC "502_ALM_ANALOG_IDB PIT 416"."VERY HIGH LEVEL VALUE (HH)" AT %DB65.DBD34, 1 s
   "502_ALM_ANALOG_IDB PIT 416_HIGH LEVEL VALUE (H)" : Real = PLC "502_ALM_ANALOG_IDB PIT 416"."HIGH LEVEL VALUE (H)" AT %DB65.DBD30, 1 s
   "502_ALM_ANALOG_IDB PIT 416_LOW LEVEL VALUE (L)" : Real = PLC "502_ALM_ANALOG_IDB PIT 416"."LOW LEVEL VALUE (L)" AT %DB65.DBD26, 1 s
   "502_ALM_ANALOG_IDB PIT 416_VERY LOW LEVEL VALUE (LL)" : Real = PLC "502_ALM_ANALOG_IDB PIT 416"."VERY LOW LEVEL VALUE (LL)" AT %DB65.DBD22, 1 s
   "IDB_PIT 402_VERY HIGH LEVEL VALUE (HH)" : Real = PLC "IDB_PIT 402"."VERY HIGH LEVEL VALUE (HH)" AT %DB742.DBD34, 1 s
   "IDB_PIT 402_HIGH LEVEL VALUE (H)" : Real = PLC "IDB_PIT 402"."HIGH LEVEL VALUE (H)" AT %DB742.DBD30, 1 s
   "IDB_PIT 402_LOW LEVEL VALUE (L)" : Real = PLC "IDB_PIT 402"."LOW LEVEL VALUE (L)" AT %DB742.DBD26, 1 s
   "IDB_PIT 402_VERY LOW LEVEL VALUE (LL)" : Real = PLC "IDB_PIT 402"."VERY LOW LEVEL VALUE (LL)" AT %DB742.DBD22, 1 s
   "TIT406_ALM_ANALOG_DB74_VERY HIGH LEVEL VALUE (HH)" : Real = PLC TIT406_ALM_ANALOG_DB74."VERY HIGH LEVEL VALUE (HH)" AT %DB74.DBD34, 1 s
   "TIT406_ALM_ANALOG_DB74_HIGH LEVEL VALUE (H)" : Real = PLC TIT406_ALM_ANALOG_DB74."HIGH LEVEL VALUE (H)" AT %DB74.DBD30, 1 s
   "TIT406_ALM_ANALOG_DB74_LOW LEVEL VALUE (L)" : Real = PLC TIT406_ALM_ANALOG_DB74."LOW LEVEL VALUE (L)" AT %DB74.DBD26, 1 s
   "TIT406_ALM_ANALOG_DB74_VERY LOW LEVEL VALUE (LL)" : Real = PLC TIT406_ALM_ANALOG_DB74."VERY LOW LEVEL VALUE (LL)" AT %DB74.DBD22, 1 s
   "LIT304_ALM_ANALOG_DB71_VERY HIGH LEVEL VALUE (HH)" : Real = PLC LIT304_ALM_ANALOG_DB71."VERY HIGH LEVEL VALUE (HH)" AT %DB71.DBD34, 1 s
   "LIT304_ALM_ANALOG_DB71_HIGH LEVEL VALUE (H)" : Real = PLC LIT304_ALM_ANALOG_DB71."HIGH LEVEL VALUE (H)" AT %DB71.DBD30, 1 s
   "LIT304_ALM_ANALOG_DB71_LOW LEVEL VALUE (L)" : Real = PLC LIT304_ALM_ANALOG_DB71."LOW LEVEL VALUE (L)" AT %DB71.DBD26, 1 s
   "LIT304_ALM_ANALOG_DB71_VERY LOW LEVEL VALUE (LL)" : Real = PLC LIT304_ALM_ANALOG_DB71."VERY LOW LEVEL VALUE (LL)" AT %DB71.DBD22, 1 s
   "IDB_TIT 315_VERY HIGH LEVEL VALUE (HH)" : Real = PLC "IDB_TIT 315"."VERY HIGH LEVEL VALUE (HH)" AT %DB715.DBD34, 1 s
   "IDB_TIT 315_HIGH LEVEL VALUE (H)" : Real = PLC "IDB_TIT 315"."HIGH LEVEL VALUE (H)" AT %DB715.DBD30, 1 s
   "IDB_TIT 315_LOW LEVEL VALUE (L)" : Real = PLC "IDB_TIT 315"."LOW LEVEL VALUE (L)" AT %DB715.DBD26, 1 s
   "IDB_TIT 315_VERY LOW LEVEL VALUE (LL)" : Real = PLC "IDB_TIT 315"."VERY LOW LEVEL VALUE (LL)" AT %DB715.DBD22, 1 s
   "IDB_TIT 401_VERY HIGH LEVEL VALUE (HH)" : Real = PLC "IDB_TIT 401"."VERY HIGH LEVEL VALUE (HH)" AT %DB741.DBD34, 1 s
   "IDB_TIT 401_HIGH LEVEL VALUE (H)" : Real = PLC "IDB_TIT 401"."HIGH LEVEL VALUE (H)" AT %DB741.DBD30, 1 s
   "IDB_TIT 401_LOW LEVEL VALUE (L)" : Real = PLC "IDB_TIT 401"."LOW LEVEL VALUE (L)" AT %DB741.DBD26, 1 s
   "IDB_TIT 401_VERY LOW LEVEL VALUE (LL)" : Real = PLC "IDB_TIT 401"."VERY LOW LEVEL VALUE (LL)" AT %DB741.DBD22, 1 s
   "IDB_PIT 102_VERY HIGH LEVEL VALUE (HH)" : Real = PLC "IDB_PIT 102"."VERY HIGH LEVEL VALUE (HH)" AT %DB722.DBD34, 1 s
   "IDB_PIT 102_HIGH LEVEL VALUE (H)" : Real = PLC "IDB_PIT 102"."HIGH LEVEL VALUE (H)" AT %DB722.DBD30, 1 s
   "IDB_PIT 102_LOW LEVEL VALUE (L)" : Real = PLC "IDB_PIT 102"."LOW LEVEL VALUE (L)" AT %DB722.DBD26, 1 s
   "IDB_PIT 102_VERY LOW LEVEL VALUE (LL)" : Real = PLC "IDB_PIT 102"."VERY LOW LEVEL VALUE (LL)" AT %DB722.DBD22, 1 s
   "PIT424PORT_ALM_ANALOG_DB_VERY HIGH LEVEL VALUE (HH)" : Real = PLC PIT424PORT_ALM_ANALOG_DB."VERY HIGH LEVEL VALUE (HH)" AT %DB2070.DBD34, 1 s
   "TT426PORT_ALM_ANALOG_DB_VERY HIGH LEVEL VALUE (HH)" : Real = PLC TT426PORT_ALM_ANALOG_DB."VERY HIGH LEVEL VALUE (HH)" AT %DB2071.DBD34, 1 s
   "TT426PORT_ALM_ANALOG_DB_HIGH LEVEL VALUE (H)" : Real = PLC TT426PORT_ALM_ANALOG_DB."HIGH LEVEL VALUE (H)" AT %DB2071.DBD30, 1 s
   "TT426PORT_ALM_ANALOG_DB_LOW LEVEL VALUE (L)" : Real = PLC TT426PORT_ALM_ANALOG_DB."LOW LEVEL VALUE (L)" AT %DB2071.DBD26, 1 s
   "TT426PORT_ALM_ANALOG_DB_VERY LOW LEVEL VALUE (LL)" : Real = PLC TT426PORT_ALM_ANALOG_DB."VERY LOW LEVEL VALUE (LL)" AT %DB2071.DBD22, 1 s
   "TT426STR_ALM_ANALOG_DB_VERY HIGH LEVEL VALUE (HH)" : Real = PLC TT426STR_ALM_ANALOG_DB."VERY HIGH LEVEL VALUE (HH)" AT %DB2072.DBD34, 1 s
   "TT426STR_ALM_ANALOG_DB_HIGH LEVEL VALUE (H)" : Real = PLC TT426STR_ALM_ANALOG_DB."HIGH LEVEL VALUE (H)" AT %DB2072.DBD30, 1 s
   "TT426STR_ALM_ANALOG_DB_LOW LEVEL VALUE (L)" : Real = PLC TT426STR_ALM_ANALOG_DB."LOW LEVEL VALUE (L)" AT %DB2072.DBD26, 1 s
